(* Logix 5000 project; controller PLC_MCC1300_75F1 vendor 1 type 14 code 166 rev 32.11; software revision 32.04; part 67 of 83 *)
(* tags used below, declared in another part *)
   CM_ConveyorStackerToLine_JS1_Sync : CM_ConveyorStackerToLine;
   CONST_dDest_Cullet : DINT;
   CONST_dDest_Stk : DINT;
   CONST_rgdDestMask : DINT[32];   // Destination Mask
   Convoy_SL_DATA_NULL : UDT_Convoy_SL;
   GP_CheckIdPlatePresent : GP_CheckIdPlatePresent;
   GP_CompactConvoy : GP_CompactConvoy;
   GP_OB_InitializeMain : GP_OB_Initialize;
   GP_RampSpace : GP_RampSpace;
   Gp_SpaceConvUtilities_V1 : GP_SpaceConvUtilities_V1;
   M311 : MAC_Conveyor;
   M311_Data : UDT_Convoy_SL;
   M316_SpaceConv_Utilities : SpaceConv_Utilities;
   M316M317_OffsetBaricentre_cmm : DINT;
   M317 : MAC_Conveyor_Single;
   M317_ALM : MAC_Conveyor_ALM;
   M317_AlmTimer1 : TIMER;
   M317_AlmTimer2 : TIMER;
   M317_Data : UDT_Convoy_SL;
   M317_dSlowingSquaringQuote : DINT;
   M317_HMW : MAC_Conveyor_HMW;
   M317_M1_DR_IN_MAM : MOTION_INSTRUCTION;
   M317_SpaceConv_Utilities : SpaceConv_Utilities;
   M317_TimerAlm3 : TIMER;
   M317_TON_Load : TIMER;
   M317_xEnableTractionRecovering : BOOL;
   M317_xPlateCullet : BOOL;
   M317_xSendCulletReqActive : BOOL;
   TMP_CenterLites : BOOL;
   TMP_d : DINT;
   TMP_dConveyorNumberForZoneCleaning : DINT;
   TMP_DistanceLateralSquaringToCenter : DINT;
   TMP_dOffsetLoadUnload_cmm : DINT;
   TMP_LiteAHeadY : DINT;
   TMP_LiteATailY : DINT;
   TMP_LiteBHeadY : DINT;
   TMP_LiteBTailY : DINT;
   TMP_rgxId : DINT[10];
   TMP_SquaringPosition : DINT;
   TMP_xConveyorInvolvedInCleaning : BOOL;
   TMP_xConveyorOfStartCleaning : BOOL;
   TMP_xCulletPresent : BOOL;
   TMP_xEnableLoadUnload : BOOL;
   TMP_xEnableZoneCleaning : BOOL;
   TMP_xLiteThisDestPresent : BOOL;
   x316PortraitMode : BOOL;
   xAlwaysOFF : BOOL;
   xAlwaysON : BOOL;
   Z402 : MAC_Zone;
   Z402_HMR : MAC_Zone_HMR;
   Z402_HMW : MAC_Zone_HMW;
   Z402S_INPUT_xSafetyAreaPopup : BOOL;
   Z402S_INPUT_xSafetyAreaRotator : BOOL;
(* MainProgram, continued *)

   32: XIC(Z402.ST_xEnableControlError)XIC(Z402S_INPUT_xSafetyAreaRotator)[XIC(M317.INPUT_xDriveInhibit_M4) ,XIC(M317.OUTPUT_xDriveEnable_M4) XIO(M317.INPUT_xDriveReady_M4) ][XIO(M317.TmON[14].DN) TON(M317.TmON[14],?,?) ,XIC(M317.TmON[14].DN) OTL(M317_ALM.rgxStoppingFault_M[0].30) ];
   33: XIC(Z402.ST_xEnableControlError)[XIC(M317.ST_xOutputEnable) [XIC(M317.PH_x.24) ,XIC(M317.PH_x.26) ] XIO(M317.tmON_AuxFunction6.DN) TON(M317.tmON_AuxFunction6,?,?) ,XIC(M317.tmON_AuxFunction6.DN) [OTL(M317_ALM.rgxWarning[0].21) ,OTL(M317.ST_xPhaseError) ] ];
   34: XIC(M317.ST_xEnableControlError)[[XIC(M317.PH_x.0) ,XIC(M317.PH_x.4) ] XIO(M317.INPUT_xLowPositionPopup_1) ,[XIC(M317.PH_x.24) XIO(M317_xEnableTractionRecovering) ,XIC(M317.PH_x.26) ,XIC(M317.PH_x.28) ] XIO(M317.INPUT_xHighPositionPopup_1) ]OTL(M317_ALM.rgxStoppingFault[0].5);
   35: XIC(M317.ST_xEnableControlError)[[XIC(M317.PH_x.0) ,XIC(M317.PH_x.4) ] XIO(M317.INPUT_xLowPositionPopup_2) ,[XIC(M317.PH_x.24) XIO(M317_xEnableTractionRecovering) ,XIC(M317.PH_x.26) ,XIC(M317.PH_x.28) ] XIO(M317.INPUT_xHighPositionPopup_2) ]OTL(M317_ALM.rgxStoppingFault[0].6);
   // Timeout rise/descent popup
   36: XIC(M317.ST_xEnableControlError)[XIC(M317.OUTPUT_xRisePopup_1) XIO(M317.INPUT_xHighPositionPopup_1) ,XIC(M317.OUTPUT_xDescentPopup_1) XIO(M317.INPUT_xLowPositionPopup_1) ,[XIC(M317.OUTPUT_xRisePopup_1) ,XIC(M317.OUTPUT_xDescentPopup_1) ] XIO(M317.INPUT_xFeedBackLiftingFrame_1) ,XIO(M317.OUTPUT_xRisePopup_1) XIO(M317.OUTPUT_xDescentPopup_1) XIC(M317.INPUT_xFeedBackLiftingFrame_1) ][XIO(M317_AlmTimer1.DN) TON(M317_AlmTimer1,?,?) ,XIC(M317_AlmTimer1.DN) OTL(M317_ALM.rgxStoppingFault[0].13) ];
   // Timeout rise/descent popup
   37: XIC(M317.ST_xEnableControlError)[XIC(M317.OUTPUT_xRisePopup_2) XIO(M317.INPUT_xHighPositionPopup_2) ,XIC(M317.OUTPUT_xDescentPopup_2) XIO(M317.INPUT_xLowPositionPopup_2) ,[XIC(M317.OUTPUT_xRisePopup_2) ,XIC(M317.OUTPUT_xDescentPopup_2) ] XIO(M317.INPUT_xFeedBackLiftingFrame_2) ,XIO(M317.OUTPUT_xRisePopup_2) XIO(M317.OUTPUT_xDescentPopup_2) XIC(M317.INPUT_xFeedBackLiftingFrame_2) ][XIO(M317_AlmTimer2.DN) TON(M317_AlmTimer2,?,?) ,XIC(M317_AlmTimer2.DN) OTL(M317_ALM.rgxStoppingFault[0].14) ];
   38: XIC(M317.ST_xEnableControlError)XIO(M317.INPUT_xProtectionLiftingFrame_1)OTL(M317_ALM.rgxStoppingFault[0].21);
   39: XIC(M317.ST_xEnableControlError)XIO(M317.INPUT_xProtectionLiftingFrame_2)OTL(M317_ALM.rgxStoppingFault[0].22);
   // Timeout feedback ventilation
   40: XIC(M317.ST_xEnableControlError)[XIC(M317.OUTPUT_xFunCommand_1) XIO(M317.INPUT_xFeedbackVentilation_1) ,XIO(M317.OUTPUT_xFunCommand_1) XIC(M317.INPUT_xFeedbackVentilation_1) ][XIO(M317.tmON_AuxFunction7.DN) TON(M317.tmON_AuxFunction7,?,?) ,XIC(M317.tmON_AuxFunction7.DN) OTL(M317_ALM.rgxWarning_M[0].0) ];
   // protection ventilation
   41: XIC(xAlwaysOFF)XIC(M317.ST_xEnableControlError)XIO(M317.INPUT_xProtectionFun_1)OTL(M317_ALM.rgxWarning_M[0].1);
   // Error position frontal squaring
   42: XIC(M317.ST_xEnableControlError)XIC(M317.ST_xOutputEnable)[XIO(M317.OUTPUT_xRiseSquaring_1) XIO(M317.INPUT_xLowPositionSquaring_1) ,XIC(M317.OUTPUT_xRiseSquaring_1) XIO(M317.INPUT_xHighPositionSquaring_1) ]XIO(M317.TmON[0].DN)[TON(M317.TmON[0],?,?) ,XIC(M317.TmON[0].DN) OTL(M317_ALM.rgxStoppingFault[0].10) ];
   // Timeout rise/descent frontal squaring
   43: XIC(M317.ST_xEnableControlError)[XIC(xAlwaysOFF) XIO(M317.INPUT_xHighPositionSquaring_1) ,XIC(M317.PH_x.8) XIO(M317.INPUT_xLowPositionSquaring_1) ][XIO(M317_TimerAlm3.DN) TON(M317_TimerAlm3,?,?) ,XIC(M317_TimerAlm3.DN) OTL(M317_ALM.rgxStoppingFault[0].11) ];
   // Timeout frontal squaring
   44: XIC(M317.ST_xEnableControlError)XIC(M317.ST_xOutputEnable)XIC(M317.PH_x.4)[XIO(M317.tmON_AuxFunction8.DN) TON(M317.tmON_AuxFunction8,?,?) ,XIC(M317.tmON_AuxFunction8.DN) [OTL(M317_ALM.rgxWarning[0].25) ,OTL(M317.ST_xPhaseError) ] ];
   // Timeout lateral squaring
   45: XIC(M317.ST_xEnableControlError)XIC(M317.ST_xOutputEnable)XIC(M317.PH_x.28)[XIO(M317.tmON_AuxFunction9.DN) TON(M317.tmON_AuxFunction9,?,?) ,XIC(M317.tmON_AuxFunction9.DN) [OTL(M317_ALM.rgxWarning[0].26) ,OTL(M317.ST_xPhaseError) ] ];
   // #####_CUMULATIVE ALARM_#####
   46: NOP();
   47: [NEQ(M317_ALM.rgxStoppingFault[0],0) ,NEQ(M317_ALM.rgxStoppingFault_M[0],0) ,NEQ(M317_ALM.rgxStoppingFault_M[1],0) ]OTE(M317.ST_xStopMachineFault);
   48: [NEQ(M317_ALM.rgxFault[0],0) ,NEQ(M317_ALM.rgxFault_M[0],0) ,NEQ(M317_ALM.rgxFault_M[1],0) ]OTE(M317.ST_xStopNextCycleFault);
END_ROUTINE

ROUTINE M317_Logic   (* ladder *)
   // #####_COSTANTS_#####
   0: [MOV(4050,TMP_dConveyorNumberForZoneCleaning) MOV(50000,TMP_dOffsetLoadUnload_cmm) MOV(500,M317_SpaceConv_Utilities.CONST_dPresetFeedbackTime_ms) OTL(TMP_xEnableLoadUnload) OTU(TMP_xEnableZoneCleaning) OTL(M317_xEnableTractionRecovering) MOV(400000,M317_SpaceConv_Utilities.CONST_dConveyorLength_cmm) MOV(775000,M317_SpaceConv_Utilities.CONST_dConveyorWidth_cmm) [GRT(Z402_HMR.dLineSpeed_mm_min,50000) XIO(M317_Data.rgtCap[0].rgxRequest.1) SUB(M317_SpaceConv_Utilities.CONST_dConveyorLength_cmm,-10000,TMP_SquaringPosition) ,LEQ(Z402_HMR.dLineSpeed_mm_min,50000) XIO(M317_Data.rgtCap[0].rgxRequest.1) SUB(M317_SpaceConv_Utilities.CONST_dConveyorLength_cmm,0,TMP_SquaringPosition) ,XIC(M317_Data.rgtCap[0].rgxRequest.1) [GRT(Z402_HMR.dLineSpeed_mm_min,50000) SUB(M317_SpaceConv_Utilities.CONST_dConveyorLength_cmm,-38000,TMP_SquaringPosition) ,LEQ(Z402_HMR.dLineSpeed_mm_min,50000) SUB(M317_SpaceConv_Utilities.CONST_dConveyorLength_cmm,-38000,TMP_SquaringPosition) ] ] ADD(TMP_SquaringPosition,M317_HMW.dParam_3_cmm,TMP_SquaringPosition) SUB(TMP_SquaringPosition,M317.AUX_dAccSpace_cmm,M317.AUX_dPresetStopLoad_cmm) ADD(M317_SpaceConv_Utilities.CONST_dConveyorLength_cmm,M317.AUX_dDecSpace_cmm,M317.AUX_dPresetStopUnload_cmm) MOV(1.2,M317_SpaceConv_Utilities.CONST_rAcceleration_ms2) MOV(1.2,M317_SpaceConv_Utilities.CONST_rDeceleration_ms2) DIV(M317_SpaceConv_Utilities.CONST_dConveyorWidth_cmm,2,TMP_DistanceLateralSquaringToCenter) MOV(388000,TMP_DistanceLateralSquaringToCenter) ,[XIC(M317.PH_x.0) [MOV(1,M317_SpaceConv_Utilities.CONST_dSyncMode) ,MOV(0,M317_SpaceConv_Utilities.CONST_dSyncroPhPosition_cmm) ,MOV(100000,M317_SpaceConv_Utilities.CONST_dSyncroPhWindow_cmm) ] ,XIC(M317.PH_x.10) [MOV(1,M317_SpaceConv_Utilities.CONST_dSyncMode) ,MOV(70000,M317_SpaceConv_Utilities.CONST_dSyncroPhPosition_cmm) ,MOV(300000,M317_SpaceConv_Utilities.CONST_dSyncroPhWindow_cmm) ] ] ];
   // #####_MATCH_#####
   1: NOP();
   // Conveyor Cleaning
   2: XIC(TMP_xEnableZoneCleaning)XIC(Z402.ST_xCleaningAccepted)GRT(Z402_HMW.dCleaningSelection,0)[EQU(Z402_HMW.dCleaningSelection,TMP_dConveyorNumberForZoneCleaning) OTE(TMP_xConveyorOfStartCleaning) ,GEQ(Z402_HMW.dCleaningSelection,TMP_dConveyorNumberForZoneCleaning) OTE(TMP_xConveyorInvolvedInCleaning) ];
   // Enable control error
   3: XIC(Z402.ST_xEnableControlError)OTE(M317.ST_xEnableControlError);
   // Mode 7 - Offsett for load/unload Simultaney
   4: XIC(M317.PH_x.8)MOV(M317.AUX_dPresetStopLoad_cmm,M317_SpaceConv_Utilities.ST_dStopLoadForseen_cmm)MOV(TMP_dOffsetLoadUnload_cmm,M317_SpaceConv_Utilities.CONF_MD7_dOffset_cmm)GP_SpaceConvUtilities_V1(Gp_SpaceConvUtilities_V1,M317_SpaceConv_Utilities,M316_SpaceConv_Utilities,M317_SpaceConv_Utilities,7);
   5: XIC(x316PortraitMode)OTU(M317_xEnableTractionRecovering);
   // Lateral position lites (referenced to baricenter, direction OpSide -> OppositeOpSide)
   6: [CPT(TMP_LiteATailY,M317_Data.rgtCap[0].rgtLite[0].dBarycenter_cmm - (M317_Data.rgtCap[0].rgtLite[0].dWidth_cmm / 2)) ,CPT(TMP_LiteAHeadY,M317_Data.rgtCap[0].rgtLite[0].dBarycenter_cmm + (M317_Data.rgtCap[0].rgtLite[0].dWidth_cmm / 2)) ,CPT(TMP_LiteBTailY,M317_Data.rgtCap[0].rgtLite[1].dBarycenter_cmm - (M317_Data.rgtCap[0].rgtLite[1].dWidth_cmm / 2)) ,CPT(TMP_LiteBHeadY,M317_Data.rgtCap[0].rgtLite[1].dBarycenter_cmm + (M317_Data.rgtCap[0].rgtLite[1].dWidth_cmm / 2)) ];
   // #####_ALARMS_#####
   7: NOP();
   // Call Alarm Routine
   8: JSR(M317_Alarm,0);
   // #####_HMI_LOGICS_#####
   9: NOP();
   // Condition ok for Cleaning
   10: [XIO(TMP_xEnableZoneCleaning) ,XIC(TMP_xEnableZoneCleaning) XIC(M317.ST_xOutputEnable) [XIO(TMP_xConveyorOfStartCleaning) ,XIC(M317.PH_x.0) ,XIO(M317.PH_x.8) ] ]OTE(M317.ST_xCleaningConditionOK);
   // Cleaning Accepted
   11: [[XIC(M317_HMW.xStopLocalCleaningRequest) ,XIC(Z402_HMW.xStopCleanZoneRequest) ] OTU(M317_HMW.xStopLocalCleaningRequest) OTU(M317_HMW.xLocalCleaningRequest) ,[XIC(M317_HMW.xLocalCleaningRequest) ,XIC(Z402.ST_xCleaningAccepted) ] [XIC(M317.ST_xCleaningConditionOK) ,XIC(M317.ST_xCleaningAccepted) ] OTE(M317.ST_xCleaningAccepted) ];
   // Manual Mode Enabled
   12: XIO(M317_SpaceConv_Utilities.ST_xFeedbackRotation)[XIC(M317_HMW.xEnableDisableManualCommand) XIC(M317.ST_xConditionOKStopCycle) OTL(M317.ST_xManualMode) ,XIO(M317_HMW.xEnableDisableManualCommand) OTU(M317.ST_xManualMode) ];
   // Virtual door enabled
   13: XIC(M317_HMW.xEnableDisableVirtualDoor)OTE(M317.ST_xVirtualDoorEnabled);
   // Clear manual command
   14: XIO(M317.ST_xManualMode)MOV(0,M317_HMW.rgxMan);
   // #####_STATUSES_#####
   15: NOP();
   // Syncro  -  OS Syncro Photocell
   16: XIC(xAlwaysON)[[XIO(M317.PH_x.10) [XIC(M317.INPUT_xSyncroPhotocell_1) ,XIC(M317.INPUT_xSyncroPhotocell_2) ] ,XIC(M317.PH_x.10) [XIC(M317.INPUT_xSquaringPhotocell_1) ,XIC(M317.INPUT_xSquaringPhotocell_2) ] ] ONS(M317.OSR_xSynchroPhotocellHead) OTE(M317.OS_xSynchroPhotocellHead) GEQ(M317_SpaceConv_Utilities.CONST_dSyncMode,1) OTE(M317_SpaceConv_Utilities.ST_OS_xSynchroPhotocellHead) ,[XIO(M317.PH_x.10) XIO(M317.INPUT_xSyncroPhotocell_1) XIO(M317.INPUT_xSyncroPhotocell_2) ,XIC(M317.PH_x.10) XIO(M317.INPUT_xSquaringPhotocell_1) XIO(M317.INPUT_xSquaringPhotocell_2) ] ONS(M317.OSR_xSynchroPhotocellTail) OTE(M317.OS_xSynchroPhotocellTail) GEQ(M317_SpaceConv_Utilities.CONST_dSyncMode,2) OTE(M317_SpaceConv_Utilities.ST_OS_xSynchroPhotocellTail) ];
   17: XIC(M317_SpaceConv_Utilities.ST_OS_xSynchroPhotocellHead)XIC(M317.PH_x.0)[MOV(0,M317_SpaceConv_Utilities.CONF_MD2_MD3_dPrstPos_cmm) GP_SpaceConvUtilities_V1(Gp_SpaceConvUtilities_V1,M317_SpaceConv_Utilities,M316_SpaceConv_Utilities,M317_SpaceConv_Utilities,2) ,SUB(0,M317_Data.dLength_cmm,M317_SpaceConv_Utilities.CONF_MD2_MD3_dPrstPos_cmm) GP_SpaceConvUtilities_V1(Gp_SpaceConvUtilities_V1,M317_SpaceConv_Utilities,M316_SpaceConv_Utilities,M317_SpaceConv_Utilities,3) ];
   // Id Plate presence
   18: MOV(CONST_rgdDestMask[24],CONST_dDest_Cullet)GP_CheckIdPlatePresent(GP_CheckIdPlatePresent,M317_Data,TMP_rgxId,M317.ST_xIdPlatePresence,TMP_xCulletPresent,CONST_dDest_Cullet)MOV(GP_CheckIdPlatePresent.OUT_dQtaLitesPresent,M317.AUX_dQtaLites)MOV(CONST_rgdDestMask[1],CONST_dDest_Stk)GP_CheckIdPlatePresent(GP_CheckIdPlatePresent,M317_Data,TMP_rgxId,M317.ST_xIdPlatePresence,TMP_xLiteThisDestPresent,CONST_dDest_Stk)XIC(TMP_xCulletPresent)OTE(M317_xPlateCullet);
   // Machine in Alarm
   19: [XIC(M317.ST_xStopMachineFault) ,XIC(M317.ST_xStopNextCycleFault) ,XIC(M317.ST_xStopNextCycleFault) ]OTE(M317.ST_xMachineAlarm);
   // Condition ok for stop Cycle
   20: [XIO(M317.ST_xPhasesInProgress) ,XIC(M317.PH_x.8) XIO(M317.OUTPUT_xRun_M1) XIO(M317_SpaceConv_Utilities.ST_xFeedbackRotation) ,XIC(M317.PH_x.12) XIO(M317.OUTPUT_xReverse_M1) XIO(M317_SpaceConv_Utilities.ST_xFeedbackRotation) ,XIC(M317.ST_xMachineAlarm) ,XIO(Z402.ST_xCycleON) ]OTE(M317.ST_xConditionOKStopCycle);
   // Cycle load unload simultaneous
   21: XIC(TMP_xEnableLoadUnload)XIO(M317.ST_xDisableLoadUnloadOnStop)XIO(M317.ST_xIdPlatePresence)OTE(M317.ST_xCycleLoadUnload);
   // Speed Management
   22: [XIO(M317_SpaceConv_Utilities.O_xRampInProgress) XIO(M317.ST_xManualMode) [MOV(Z402_HMR.dLineSpeed_mm_min,M317.AUX_dReqSpeed_mm_min) ,XIC(M317.PH_x.4) MOV(10000,M317.AUX_dReqSpeed_mm_min) ] ,XIC(M317.ST_xManualMode) MOV(Z402_HMW.dManualSpeed_mm_min,M317.AUX_dReqSpeed_mm_min) ,NEQ(M317.AUX_dReqSpeed_mm_min,M317_SpaceConv_Utilities.ST_dRealSpeed_mm_min) OTE(M317.OS_xChangeSpeed) ];
   // Ramp Management
   23: GP_RampSpace(GP_RampSpace,M317_SpaceConv_Utilities.CONST_rAcceleration_ms2,M317_SpaceConv_Utilities.CONST_rDeceleration_ms2,M317_SpaceConv_Utilities.ST_dRealSpeed_mm_min,M317.AUX_dAccSpace_cmm,M317.AUX_dDecSpace_cmm);
   // Space Convoy utilities MOD 1 for Calculate Head/Tail
   24: XIC(xAlwaysON)[[XIC(M317.OUTPUT_xRun_M1) ,XIC(M317.OUTPUT_xReverse_M1) ] XIO(M317.ST_xManualMode) OTE(M317_SpaceConv_Utilities.CONF_MD1_xRun) ,XIC(M317.OUTPUT_xReverse_M1) XIC(xAlwaysOFF) XIO(M317.ST_xManualMode) OTE(M317_SpaceConv_Utilities.CONF_MD1_xReverse) ,[XIC(M317.INPUT_xDriveFeedback_M1) ,XIC(M317_SpaceConv_Utilities.CONF_MD1_xRun) GRT(M317_SpaceConv_Utilities.O_dCountFeedbackTime_ms,0) ] OTE(M317_SpaceConv_Utilities.ST_xFeedbackRotation) ,XIC(M317.ST_xIdPlatePresence) OTE(M317_SpaceConv_Utilities.CONF_MD1_xHeadTracking) ,XIC(M317.ST_xPlatePresence) OTE(M317_SpaceConv_Utilities.CONF_MD1_xTailTracking) ,MOV(GP_OB_InitializeMain.OUT_dExecutionTime_ms,M317_SpaceConv_Utilities.CONF_MD1_dScan_ms) GP_SpaceConvUtilities_V1(Gp_SpaceConvUtilities_V1,M317_SpaceConv_Utilities,M316_SpaceConv_Utilities,M317_SpaceConv_Utilities,1) ];
   // Output Enable
   25: XIC(Z402.ST_xCycleON)XIO(M317.ST_xManualMode)XIO(M317.ST_xStopMachineFault)[XIO(M317.ST_xPlatePassageUpstream_FW) XIO(M317.ST_xPlatePassageUpstream_BKW) ,XIC(M317.ST_xPlatePassageUpstream_FW) XIC(M311.ST_xOutputEnable) ,XIC(M317.ST_xPlatePassageUpstream_BKW) XIC(CM_ConveyorStackerToLine_JS1_Sync.xOutputEnable) ]XIC(Z402S_INPUT_xSafetyAreaPopup)OTE(M317.ST_xOutputEnable);
   26: XIC(TMP_xLiteThisDestPresent)OTL(M317_xSendCulletReqActive);
   27: XIO(TMP_xLiteThisDestPresent)OTU(M317_xSendCulletReqActive);
   // #####_WORKING_FLAGS_#####
   28: NOP();
   // Frontal squaring request
   29: XIC(M317.OS_xLoad_FW)[NEQ(M317_Data.rgtCap[0].rgtLite[0].dID,0) GEQ(M317_Data.rgtCap[0].rgtLite[0].dWidth_cmm,M317_Data.rgtCap[0].dLength_cmm) ,NEQ(M317_Data.rgtCap[0].rgtLite[1].dID,0) GEQ(M317_Data.rgtCap[0].rgtLite[1].dWidth_cmm,M317_Data.rgtCap[0].dLength_cmm) ]XIO(TMP_xCulletPresent)OTL(M317_Data.rgtCap[0].rgxRequest.0);
   // Lateral squaring request
   30: XIC(M317.OS_xLoad_FW)[NEQ(M317_Data.rgtCap[0].rgtLite[0].dID,0) GRT(M317_Data.rgtCap[0].dLength_cmm,M317_Data.rgtCap[0].rgtLite[0].dWidth_cmm) ,NEQ(M317_Data.rgtCap[0].rgtLite[1].dID,0) GRT(M317_Data.rgtCap[0].dLength_cmm,M317_Data.rgtCap[0].rgtLite[1].dWidth_cmm) ]XIO(TMP_xCulletPresent)OTL(M317_Data.rgtCap[0].rgxRequest.1);
   // Adjust position for stacker
   31: XIC(M317.ST_xIdPlatePresence)XIO(TMP_xCulletPresent)[XIC(M317_Data.rgtCap[0].rgxDone.0) ,XIC(M317_Data.rgtCap[0].rgxDone.1) ][[NEQ(M317_Data.rgtCap[0].rgtLite[0].dID,0) NEQ(M317_Data.rgtCap[0].rgtLite[0].dBarycenter_cmm,0) ,NEQ(M317_Data.rgtCap[0].rgtLite[1].dID,0) NEQ(M317_Data.rgtCap[0].rgtLite[1].dBarycenter_cmm,0) ] ,NEQ(M317_Data.rgtCap[0].rgtLite[0].dID,0) NEQ(M317_Data.rgtCap[0].rgtLite[1].dID,0) [GRT(TMP_LiteAHeadY,0) ,LES(TMP_LiteBTailY,0) ] OTE(TMP_CenterLites) ]OTL(M317_Data.rgtCap[0].rgxRequest.2);
   // #####_LOGICS_#####
   32: NOP();
   // Phase of load
   33: XIC(M311.OS_xUnload_FW)[OTL(M317.PH_x.0) ,OTU(M317_SpaceConv_Utilities.O_xPlateSynchronized) ,OTU(M317.ST_xDisableLoadUnloadOnStop) ,OTE(M317.OS_xLoad_FW) ,XIC(M311.OS_xUnload_FW) COP(M311_Data,M317_Data,1) CPT(M317_Data.rgtCap[0].rgtLite[0].dBarycenter_cmm,M317_Data.rgtCap[0].rgtLite[0].dBarycenter_cmm - M316M317_OffsetBaricentre_cmm) FLL(0,M311_Data,1) GP_CompactConvoy(GP_CompactConvoy,M317_Data,Convoy_SL_DATA_NULL) ,GP_SpaceConvUtilities_V1(Gp_SpaceConvUtilities_V1,M317_SpaceConv_Utilities,M316_SpaceConv_Utilities,M317_SpaceConv_Utilities,5) ,NEQ(M317_Data.rgtCap[0].rgtLite[0].dID,0) NEQ(M317_Data.rgtCap[0].rgtLite[1].dID,0) MOV(2,M317_Data.rgtCap[0].dNumLites) MOV(25000,M317_Data.rgtCap[0].dGap_cmm) CPT(M317_Data.rgtCap[0].dWidth_cmm,(M317_Data.rgtCap[0].dWidth_cmm * 2) + M317_Data.rgtCap[0].dGap_cmm) ];
   // Request positioning
   34: NOP();
   // Syncro  -  Space Convoy utilities MOD 4
   35: GRT(M317_SpaceConv_Utilities.CONST_dSyncMode,0)[XIC(M317.PH_x.0) XIO(M317.PH_x.8) ,XIC(M317.PH_x.0) XIC(M317.PH_x.8) ADD(M317_SpaceConv_Utilities.CONST_dSyncroPhPosition_cmm,TMP_dOffsetLoadUnload_cmm,TMP_d) GRT(M317_SpaceConv_Utilities.O_dTailPosition_cmm,TMP_d) ][MOV(M317_Data.dLength_cmm,M317_SpaceConv_Utilities.CONF_MD4_MD6_dLength_cmm) ,GP_SpaceConvUtilities_V1(Gp_SpaceConvUtilities_V1,M317_SpaceConv_Utilities,M316_SpaceConv_Utilities,M317_SpaceConv_Utilities,4) ];
   36: XIC(M317.PH_x.0)XIC(M317.ST_xOutputEnable)[XIC(M317.OUTPUT_xRun_M1) ,XIC(M317.OUTPUT_xRun_M2) ]SUB(M317_SpaceConv_Utilities.CONST_dConveyorLength_cmm,M317.AUX_dAccSpace_cmm,M317_dSlowingSquaringQuote)DIV(Z402_HMR.dLineSpeed_mm_min,6000,TMP_d)DIV(M317_dSlowingSquaringQuote,TMP_d,TMP_d)DIV(TMP_d,10,M317_TON_Load.PRE)TON(M317_TON_Load,?,?);
   // End load Phase
   37: XIC(M317.PH_x.0)[XIO(M317_Data.tFlag.tConveyor.xReqStop) GRT(M317_SpaceConv_Utilities.O_dHeadPosition_cmm,M317.AUX_dPresetStopLoad_cmm) XIO(M317.INPUT_xSyncroPhotocell_1) ,XIC(M317_Data.tFlag.tConveyor.xReqStop) [XIC(M317.OUTPUT_xPositioning_M1) XIC(M317_M1_DR_IN_MAM.PC) ,XIC(M317.ST_xPhaseError) ] ][OTE(M317.PH_x.7) ,OTU(M317.PH_x.0) ,OTL(M317.ST_xPlatePresence) ];
   // End positiong
   38: XIC(M317.PH_x.7)XIC(M317_Data.tFlag.tConveyor.xReqStop)XIC(M317.OUTPUT_xPositioning_M1)XIC(M317_M1_DR_IN_MAM.PC)[OTU(M317_Data.tFlag.tConveyor.xReqStop) ,OTL(M317_Data.tFlag.tConveyor.xReqStopEndConveyor) ,CPT(M317_SpaceConv_Utilities.CONF_MD2_MD3_dPrstPos_cmm,TMP_SquaringPosition) GP_SpaceConvUtilities_V1(Gp_SpaceConvUtilities_V1,M317_SpaceConv_Utilities,M316_SpaceConv_Utilities,M317_SpaceConv_Utilities,2) ];
